// TIA Portal project "TestEssProtoFreia" (V13) (continued)
REGION Network 9: Reset SND_BUSY flag when completed without errors
   RUNG wire#powerrail
      Contact( "SND_DONE(1)" )
      Contact( "SND_BUSY(1)" )
      R_Coil( "SND_BUSY(1)" )
   END_RUNG
   // the same network as SCL:
   IF "SND_DONE(1)" AND "SND_BUSY(1)" THEN "SND_BUSY(1)" := FALSE; END_IF;
END_REGION

REGION Network 10 (STL): Reset SND_BUSY flag and save the status when returned error
         AN    "SND_DONE(1)";
         A     "SND_ERR(1)";
         JNB   ex2;
         R     "SND_BUSY(1)";
         L     "SEND_status(1)";
         T     "SND_STAT_SAVE(1)";
   ex2:  NOP   0;
END_REGION
END_FUNCTION

FUNCTION "Recv_from_Epics" : Void   // FC31, STL
{ S7_Optimized_Access := 'FALSE' }
VERSION : 0.1
BEGIN

REGION Network 1: Get data from Epics (channel 1)
         CALL  AG_RECV
         ( ID     := 1,
           LADDR  := w#16#400,
           RECV   := P#DB101.DBX0.0 BYTE 1000,
           NDR    := "RCV_NDR",
           ERROR  := "RCV_ERR",
           STATUS := "RECV_status",
           LEN    := "RECV_len"
         );
         AN    "RCV_NDR";
         O     "RCV_ERR";
         JC    out;
         CALL  "Cmds_from_Epics";
         BE;
   out:  AN    "RCV_ERR";
         JC    _001;
         L     "RECV_status";
         T     "RCV_STAT_SAVE";
   _001: NOP   0;
END_REGION

REGION Network 2: Get data from Epics (channel 2)
         CALL  AG_RECV
         ( ID     := 2,
           LADDR  := w#16#400,
           RECV   := P#DB105.DBX0.0 BYTE 250,
           NDR    := "RCV_NDR(1)",
           ERROR  := "RCV_ERR(1)",
           STATUS := "RECV_status(1)",
           LEN    := "RECV_len(1)"
         );
         AN    "RCV_NDR(1)";
         O     "RCV_ERR(1)";
         JC    out2;
         CALL  "Data_from_IOC";
         BE;
   out2: AN    "RCV_ERR(1)";
         JC    _002;
         L     "RECV_status(1)";
         T     "RCV_STAT_SAVE(1)";
   _002: NOP   0;
END_REGION
END_FUNCTION

FUNCTION "Send_Epics_data" : Void   // FC32, STL
{ S7_Optimized_Access := 'FALSE' }
VERSION : 0.1
BEGIN

REGION Network 2: Update the Local/remote status
         A     "LocalMode";
         =     "PLC_to_Epics".sLocal;
END_REGION

REGION Network 3: CV01
         L     "CV01_HMI_VAL";
         T     "PLC_to_Epics".CV01.sSetV;
         L     "Tag_7";
         T     "PLC_to_Epics".CV01.sRdV;

         AN    "CV01_ManAuto";
         =     "PLC_to_Epics".CV01.sAuto;
END_REGION

REGION Network 4: CV02
         L     "CV02_HMI_VAL";
         T     "PLC_to_Epics".CV02.sSetV;
         L     "Tag_8";
         T     "PLC_to_Epics".CV02.sRdV;

         AN    "CV02_ManAuto";
         =     "PLC_to_Epics".CV02.sAuto;
END_REGION

REGION Network 5: CV03
         L     "CV03_HMI_VAL";
         T     "PLC_to_Epics".CV03.sSetV;
         L     "Tag_9";
         T     "PLC_to_Epics".CV03.sRdV;

         AN    "CV03_ManAuto";
         =     "PLC_to_Epics".CV03.sAuto;
END_REGION

REGION Network 6: CV04
         L     "CV04_HMI_VAL";
         T     "PLC_to_Epics".CV04.sSetV;
         L     "Tag_10";
         T     "PLC_to_Epics".CV04.sRdV;

         AN    "CV04_ManAuto";
         =     "PLC_to_Epics".CV04.sAuto;
END_REGION

REGION Network 7: CV05
         L     "CV05_HMI_VAL";
         T     "PLC_to_Epics".CV05.sSetV;
         L     "Tag_11";
         T     "PLC_to_Epics".CV05.sRdV;

   //      AN    "CV05_ManAuto"
   //      =     "PLC_to_Epics".CV05.sAuto
END_REGION

REGION Network 8: CV07
         L     "CV07_HMI_VAL";
         T     "PLC_to_Epics".CV07.sSetV;
         L     "Tag_12";
         T     "PLC_to_Epics".CV07.sRdV;

         AN    "CV07_ManAuto";
         =     "PLC_to_Epics".CV07.sAuto;
END_REGION

REGION Network 9: CV60
         L     "CV60_HMI_VAL";
         T     "PLC_to_Epics".CV60.sSetV;
         L     "Tag_13";
         T     "PLC_to_Epics".CV60.sRdV;

         AN    "CV60_ManAuto";
         =     "PLC_to_Epics".CV60.sAuto;
END_REGION

REGION Network 10: CV61
         L     "CV61_HMI_VAL";
         T     "PLC_to_Epics".CV61.sSetV;
         L     "Tag_14";
         T     "PLC_to_Epics".CV61.sRdV;

         AN    "CV61_ManAuto";
         =     "PLC_to_Epics".CV61.sAuto;
END_REGION

REGION Network 11: CV62
         L     "CV62_HMI_VAL";
         T     "PLC_to_Epics".CV62.sSetV;
         L     "Tag_15";
         T     "PLC_to_Epics".CV62.sRdV;

   //      AN    "CV62_ManAuto"
   //      =     "PLC_to_Epics".CV62.sAuto
END_REGION

REGION Network 12: CV550
   //      L     "Tag_14"
   //      T     "PLC_to_Epics".CV550.sRdV

         AN    "ASCOenManuel";
         =     "PLC_to_Epics".CV550.sAuto;
         =     "Data_fo_HNOSS".RegOnMKS2;
END_REGION

REGION Network 13: spare - VB chan 7
         A     "voie 7 chaufferette BV";
         =     "PLC_to_Epics"."spare-VB-7".sHtrOn;
END_REGION

REGION Network 14: spare - VB chan 8
         A     "voie 8 chaufferette BV";
         =     "PLC_to_Epics"."spare-VB-8".sHtrOn;
END_REGION

REGION Network 15: spare VB chan 9
         A     "voie 9 chaufferette BV";
         =     "PLC_to_Epics"."spare-VB-9".sHtrOn;
END_REGION

REGION Network 16: spare - VB chan 10
         A     "voie 10  chaufferette BV";
         =     "PLC_to_Epics"."spare-VB-10".sHtrOn;
END_REGION

REGION Network 17: spare - VB chan 11
         A     "voie 11 chaufferette BV";
         =     "PLC_to_Epics"."spare-VB-11".sHtrOn;
END_REGION

REGION Network 18: EH901-902 CM chan 1
         A     "voie 1 chaufferette CM";
         =     "PLC_to_Epics".EH01.sHtrOn;
END_REGION

REGION Network 19: EH913-914 CM channel 4
         A     "voie 4 chaufferette CM";
         =     "PLC_to_Epics".EH20.sHtrOn;
END_REGION

REGION Network 20: EH933-934 - CM chan 5
         A     "voie 5 chaufferette CM";
         =     "PLC_to_Epics"."spare-CM-5".sHtrOn;
END_REGION

REGION Network 21: EH921 - CM chan 6
         A     "voie 6 chaufferette CM";
         =     "PLC_to_Epics"."spare-CM-6".sHtrOn;
END_REGION

REGION Network 22: EH931-932 - CM chan 7
         A     "voie 7 chaufferette CM";
         =     "PLC_to_Epics"."spare-CM-7".sHtrOn;
END_REGION

REGION Network 23: EH915-916 - CM chan 8
         A     "voie 8 chaufferette CM";
         =     "PLC_to_Epics"."spare-CM-8".sHtrOn;
END_REGION

REGION Network 24: EH937-938 - CM chan 10
         A     "voie 10 chaufferette CM";
         =     "PLC_to_Epics"."spare-CM-10".sHtrOn;
END_REGION

REGION Network 25: EH935-936 - CM chan 12
         A     "voie 12 chaufferette CM";
         =     "PLC_to_Epics"."spare-CM-12".sHtrOn;
END_REGION

REGION Network 26: Status bits
         A     "Graph/manuelle";
         =     "PLC_to_Epics".sManual;
         A     "ErreurSupervision";
         =     "PLC_to_Epics".sGrafcetERR;
         A     "Etat initial";
         =     "PLC_to_Epics".sGS1;
         A     "EtatCdtCryo";
         =     "PLC_to_Epics".sGS2;
         A     "EtatAttMef";
         =     "PLC_to_Epics".sGS3;
         A     "EtatMEFazote";
         =     "PLC_to_Epics".sGS4;
         A     "EtatMEFhelium";
         =     "PLC_to_Epics".sGS5;
         A     "EtatMode4k";
         =     "PLC_to_Epics".sGS6;
         A     "EtatModeStandBy";
         =     "PLC_to_Epics".sGS7;
         A     "EtatMode2K";
         =     "PLC_to_Epics".sGS8;
         A     "Etatrechauffage";
         =     "PLC_to_Epics".sGS10;
         A     "conditionTempMEFheliumOK";
         =     "PLC_to_Epics".sTransTempOK;
         A     "TransMode4K";
         =     "PLC_to_Epics".sTransMode4K;
         A     "EPICS_COMM_OK";
         =     "PLC_to_Epics".EpicsCommOK;
         A     "HNOSS_COMM_OK";
         =     "PLC_to_Epics".HNOSSCommOK;
END_REGION

REGION Network 27: Real parameters read-back (LHe level PID settings)
         L     "TriggerPIDcv01";
         T     "PLC_to_Epics".TrigPID_CV01.sSetV;
         L     "TriggerPIDcv02";
         T     "PLC_to_Epics".TrigPID_CV02.sSetV;
         L     "TriggerPIDcv03";
         T     "PLC_to_Epics".TrigPID_CV03.sSetV;
         L     "LT01LevelSP2k";
         T     "PLC_to_Epics".PID_LT01_CV01_SP.sSetV;
         L     "LT01LevelSP";
         T     "PLC_to_Epics".PID_LT01_CV02_SP.sSetV;
         L     "LT03LevelSP";
         T     "PLC_to_Epics".PID_LT03_CV03_SP.sSetV;
END_REGION

REGION Network 28: Real parameters read-back (CV550l PID settings)
         L     "RéguleASCO02_SP";
         T     "PLC_to_Epics".PID_PT01_CV550_SP.sSetV;
END_REGION

REGION Network 29: Sequence steps
         L     "Data_fo_HNOSS".S4step;
         T     "PLC_to_Epics".S4step;
         L     "Data_fo_HNOSS".S5step;
         T     "PLC_to_Epics".S5step;
         L     "Data_fo_HNOSS".S6step;
         T     "PLC_to_Epics".S6step;
         L     "Data_fo_HNOSS".S7step;
         T     "PLC_to_Epics".S7step;
         L     "Data_fo_HNOSS".S8step;
         T     "PLC_to_Epics".S8step;
         L     "Data_fo_HNOSS".S9step;
         T     "PLC_to_Epics".S9step;
         L     "Data_fo_HNOSS".S10step;
         T     "PLC_to_Epics".S10step;
         L     "Data_fo_HNOSS".SXstep;
         T     "PLC_to_Epics".SXstep;
END_REGION
END_FUNCTION

FUNCTION "Cmds_from_Epics" : Void   // FC33, LAD
TITLE = Process data from Epics
{ S7_Optimized_Access := 'FALSE' }
VERSION : 0.1
   VAR_TEMP   // added for the SCL form of the ladder/FBD networks
      _w1 : Bool;
   END_VAR
BEGIN

REGION Network 1: Switch to remote mode (control from Epics)
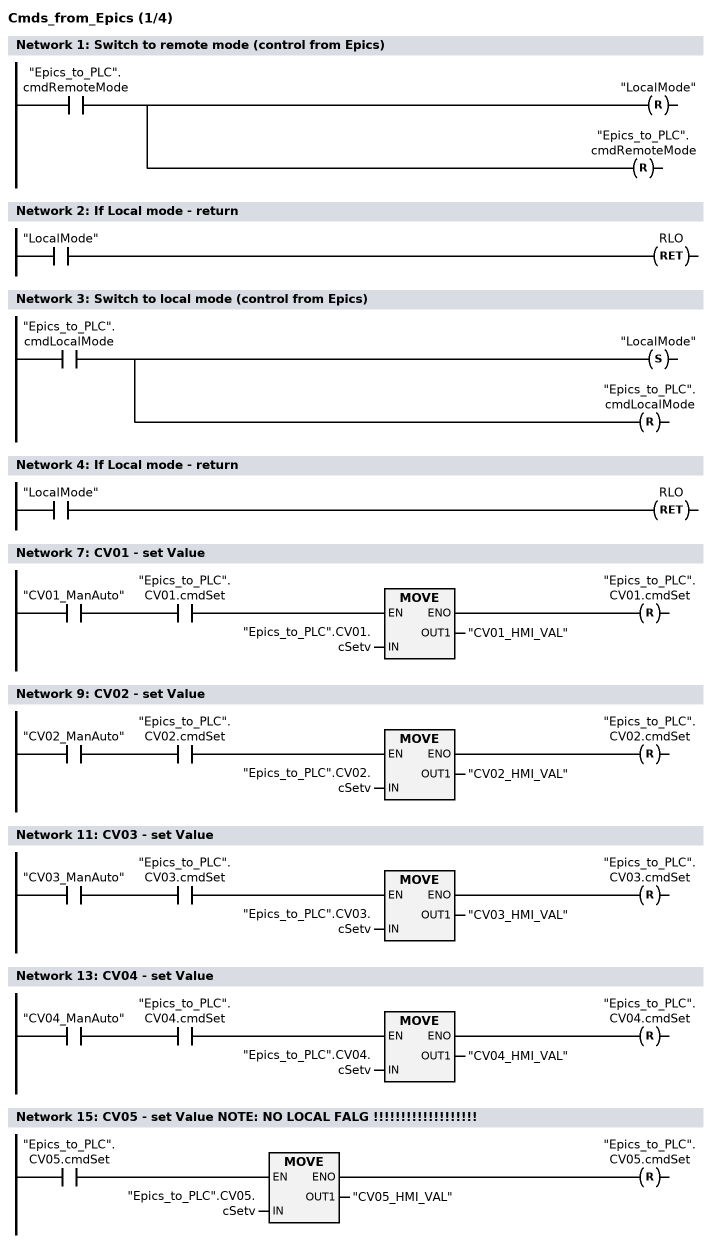
   RUNG wire#powerrail
      Contact( "Epics_to_PLC".cmdRemoteMode )
      wire#w1
      R_Coil( "LocalMode" )
   END_RUNG
   RUNG wire#w1
      R_Coil( "Epics_to_PLC".cmdRemoteMode )
   END_RUNG
   // the same network as SCL:
   IF "Epics_to_PLC".cmdRemoteMode THEN
       "LocalMode" := FALSE;
       "Epics_to_PLC".cmdRemoteMode := FALSE;
   END_IF;
END_REGION

REGION Network 2: If Local mode - return
   IF "LocalMode" THEN
       ENO := TRUE;
       RETURN;
   END_IF;
END_REGION

REGION Network 3: Switch to local mode (control from Epics)
   RUNG wire#powerrail
      Contact( "Epics_to_PLC".cmdLocalMode )
      wire#w1
      S_Coil( "LocalMode" )
   END_RUNG
   RUNG wire#w1
      R_Coil( "Epics_to_PLC".cmdLocalMode )
   END_RUNG
   // the same network as SCL:
   IF "Epics_to_PLC".cmdLocalMode THEN
       "LocalMode" := TRUE;
       "Epics_to_PLC".cmdLocalMode := FALSE;
   END_IF;
END_REGION

REGION Network 4: If Local mode - return
   IF "LocalMode" THEN
       ENO := TRUE;
       RETURN;
   END_IF;
END_REGION

REGION Network 5: Test data (copy block of data)
END_REGION

REGION Network 6 (STL): CV01 Man/Auto
         A     "Epics_to_PLC".CV01.cmdAuto;
         R     "CV01_ManAuto";
         A     "Epics_to_PLC".CV01.cmdMan;
         S     "CV01_ManAuto";
END_REGION

REGION Network 7: CV01 - set Value
   RUNG wire#powerrail
      Contact( "CV01_ManAuto" )
      Contact( "Epics_to_PLC".CV01.cmdSet )
      { S7_GenerateENO := "TRUE" } Move(in := "Epics_to_PLC".CV01.cSetv, out1 => "CV01_HMI_VAL")
      R_Coil( "Epics_to_PLC".CV01.cmdSet )
   END_RUNG
   // the same network as SCL:
   // ENO of a box is taken as its EN; it also drops when the box reports an error
   IF "CV01_ManAuto" AND "Epics_to_PLC".CV01.cmdSet THEN
       "CV01_HMI_VAL" := "Epics_to_PLC".CV01.cSetv;
       "Epics_to_PLC".CV01.cmdSet := FALSE;
   END_IF;
END_REGION

REGION Network 8 (STL): CV02 Man/Auto
         A     "Epics_to_PLC".CV02.cmdAuto;
         R     "CV02_ManAuto";
         A     "Epics_to_PLC".CV02.cmdMan;
         S     "CV02_ManAuto";
END_REGION

REGION Network 9: CV02 - set Value
   RUNG wire#powerrail
      Contact( "CV02_ManAuto" )
      Contact( "Epics_to_PLC".CV02.cmdSet )
      { S7_GenerateENO := "TRUE" } Move(in := "Epics_to_PLC".CV02.cSetv, out1 => "CV02_HMI_VAL")
      R_Coil( "Epics_to_PLC".CV02.cmdSet )
   END_RUNG
   // the same network as SCL:
   // ENO of a box is taken as its EN; it also drops when the box reports an error
   IF "CV02_ManAuto" AND "Epics_to_PLC".CV02.cmdSet THEN
       "CV02_HMI_VAL" := "Epics_to_PLC".CV02.cSetv;
       "Epics_to_PLC".CV02.cmdSet := FALSE;
   END_IF;
END_REGION

REGION Network 10 (STL): CV03 Man/Auto
         A     "Epics_to_PLC".CV03.cmdAuto;
         R     "CV03_ManAuto";
         A     "Epics_to_PLC".CV03.cmdMan;
         S     "CV03_ManAuto";
END_REGION

REGION Network 11: CV03 - set Value
   RUNG wire#powerrail
      Contact( "CV03_ManAuto" )
      Contact( "Epics_to_PLC".CV03.cmdSet )
      { S7_GenerateENO := "TRUE" } Move(in := "Epics_to_PLC".CV03.cSetv, out1 => "CV03_HMI_VAL")
      R_Coil( "Epics_to_PLC".CV03.cmdSet )
   END_RUNG
   // the same network as SCL:
   // ENO of a box is taken as its EN; it also drops when the box reports an error
   IF "CV03_ManAuto" AND "Epics_to_PLC".CV03.cmdSet THEN
       "CV03_HMI_VAL" := "Epics_to_PLC".CV03.cSetv;
       "Epics_to_PLC".CV03.cmdSet := FALSE;
   END_IF;
END_REGION

REGION Network 12 (STL): CV04 Man/Auto
         A     "Epics_to_PLC".CV04.cmdAuto;
         R     "CV04_ManAuto";
         A     "Epics_to_PLC".CV04.cmdMan;
         S     "CV04_ManAuto";
END_REGION

REGION Network 13: CV04 - set Value
   RUNG wire#powerrail
      Contact( "CV04_ManAuto" )
      Contact( "Epics_to_PLC".CV04.cmdSet )
      { S7_GenerateENO := "TRUE" } Move(in := "Epics_to_PLC".CV04.cSetv, out1 => "CV04_HMI_VAL")
      R_Coil( "Epics_to_PLC".CV04.cmdSet )
   END_RUNG
   // the same network as SCL:
   // ENO of a box is taken as its EN; it also drops when the box reports an error
   IF "CV04_ManAuto" AND "Epics_to_PLC".CV04.cmdSet THEN
       "CV04_HMI_VAL" := "Epics_to_PLC".CV04.cSetv;
       "Epics_to_PLC".CV04.cmdSet := FALSE;
   END_IF;
END_REGION

REGION Network 14: CV05 Man/Auto
END_REGION

REGION Network 15: CV05 - set Value NOTE: NO LOCAL FALG !!!!!!!!!!!!!!!!!!!
   RUNG wire#powerrail
      Contact( "Epics_to_PLC".CV05.cmdSet )
      { S7_GenerateENO := "TRUE" } Move(in := "Epics_to_PLC".CV05.cSetv, out1 => "CV05_HMI_VAL")
      R_Coil( "Epics_to_PLC".CV05.cmdSet )
   END_RUNG
   // the same network as SCL:
   // ENO of a box is taken as its EN; it also drops when the box reports an error
   IF "Epics_to_PLC".CV05.cmdSet THEN
       "CV05_HMI_VAL" := "Epics_to_PLC".CV05.cSetv;
       "Epics_to_PLC".CV05.cmdSet := FALSE;
   END_IF;
END_REGION

REGION Network 16 (STL): CV07 Man/Auto
         A     "Epics_to_PLC".CV07.cmdAuto;
         R     "CV07_ManAuto";
         A     "Epics_to_PLC".CV07.cmdMan;
         S     "CV07_ManAuto";
END_REGION

REGION Network 17: CV07 - set Value
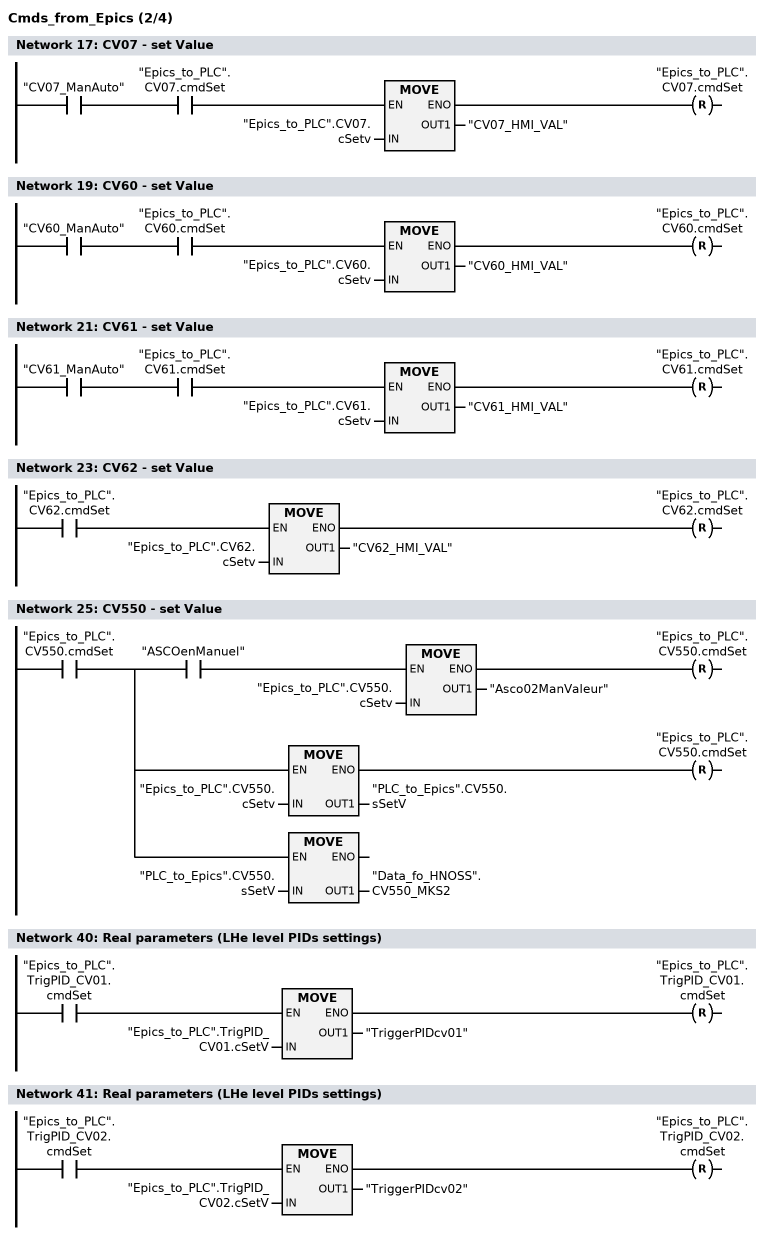
   RUNG wire#powerrail
      Contact( "CV07_ManAuto" )
      Contact( "Epics_to_PLC".CV07.cmdSet )
      { S7_GenerateENO := "TRUE" } Move(in := "Epics_to_PLC".CV07.cSetv, out1 => "CV07_HMI_VAL")
      R_Coil( "Epics_to_PLC".CV07.cmdSet )
   END_RUNG
   // the same network as SCL:
   // ENO of a box is taken as its EN; it also drops when the box reports an error
   IF "CV07_ManAuto" AND "Epics_to_PLC".CV07.cmdSet THEN
       "CV07_HMI_VAL" := "Epics_to_PLC".CV07.cSetv;
       "Epics_to_PLC".CV07.cmdSet := FALSE;
   END_IF;
END_REGION

REGION Network 18 (STL): CV60 Man/Auto
         A     "Epics_to_PLC".CV60.cmdAuto;
         R     "CV60_ManAuto";
         A     "Epics_to_PLC".CV60.cmdMan;
         S     "CV60_ManAuto";
END_REGION

REGION Network 19: CV60 - set Value
   RUNG wire#powerrail
      Contact( "CV60_ManAuto" )
      Contact( "Epics_to_PLC".CV60.cmdSet )
      { S7_GenerateENO := "TRUE" } Move(in := "Epics_to_PLC".CV60.cSetv, out1 => "CV60_HMI_VAL")
      R_Coil( "Epics_to_PLC".CV60.cmdSet )
   END_RUNG
   // the same network as SCL:
   // ENO of a box is taken as its EN; it also drops when the box reports an error
   IF "CV60_ManAuto" AND "Epics_to_PLC".CV60.cmdSet THEN
       "CV60_HMI_VAL" := "Epics_to_PLC".CV60.cSetv;
       "Epics_to_PLC".CV60.cmdSet := FALSE;
   END_IF;
END_REGION

REGION Network 20 (STL): CV61 Man/Auto
         A     "Epics_to_PLC".CV61.cmdAuto;
         R     "CV61_ManAuto";
         A     "Epics_to_PLC".CV61.cmdMan;
         S     "CV61_ManAuto";
END_REGION

REGION Network 21: CV61 - set Value
   RUNG wire#powerrail
      Contact( "CV61_ManAuto" )
      Contact( "Epics_to_PLC".CV61.cmdSet )
      { S7_GenerateENO := "TRUE" } Move(in := "Epics_to_PLC".CV61.cSetv, out1 => "CV61_HMI_VAL")
      R_Coil( "Epics_to_PLC".CV61.cmdSet )
   END_RUNG
   // the same network as SCL:
   // ENO of a box is taken as its EN; it also drops when the box reports an error
   IF "CV61_ManAuto" AND "Epics_to_PLC".CV61.cmdSet THEN
       "CV61_HMI_VAL" := "Epics_to_PLC".CV61.cSetv;
       "Epics_to_PLC".CV61.cmdSet := FALSE;
   END_IF;
END_REGION

REGION Network 22: CV62 Man/Auto
END_REGION

REGION Network 23: CV62 - set Value
   RUNG wire#powerrail
      Contact( "Epics_to_PLC".CV62.cmdSet )
      { S7_GenerateENO := "TRUE" } Move(in := "Epics_to_PLC".CV62.cSetv, out1 => "CV62_HMI_VAL")
      R_Coil( "Epics_to_PLC".CV62.cmdSet )
   END_RUNG
   // the same network as SCL:
   // ENO of a box is taken as its EN; it also drops when the box reports an error
   IF "Epics_to_PLC".CV62.cmdSet THEN
       "CV62_HMI_VAL" := "Epics_to_PLC".CV62.cSetv;
       "Epics_to_PLC".CV62.cmdSet := FALSE;
   END_IF;
END_REGION

REGION Network 24 (STL): CV550 Man/Auto
         A     "Epics_to_PLC".CV550.cmdAuto;
         R     "ASCOenManuel";
         A     "Epics_to_PLC".CV550.cmdMan;
         S     "ASCOenManuel";
END_REGION

REGION Network 25: CV550 - set Value
   RUNG wire#powerrail
      Contact( "Epics_to_PLC".CV550.cmdSet )
      wire#w1
      Contact( "ASCOenManuel" )
      { S7_GenerateENO := "TRUE" } Move(in := "Epics_to_PLC".CV550.cSetv, out1 => "Asco02ManValeur")
      R_Coil( "Epics_to_PLC".CV550.cmdSet )
   END_RUNG
   RUNG wire#w1
      { S7_GenerateENO := "TRUE" } Move(in := "Epics_to_PLC".CV550.cSetv, out1 => "PLC_to_Epics".CV550.sSetV)
      R_Coil( "Epics_to_PLC".CV550.cmdSet )
   END_RUNG
   RUNG wire#w1
      { S7_GenerateENO := "TRUE" } Move(in := "PLC_to_Epics".CV550.sSetV, out1 => "Data_fo_HNOSS".CV550_MKS2)
   END_RUNG
   // the same network as SCL:
   // ENO of a box is taken as its EN; it also drops when the box reports an error
   IF "Epics_to_PLC".CV550.cmdSet AND "ASCOenManuel" THEN
       "Asco02ManValeur" := "Epics_to_PLC".CV550.cSetv;
   END_IF;
   #_w1 := "Epics_to_PLC".CV550.cmdSet;
   IF "Epics_to_PLC".CV550.cmdSet AND "ASCOenManuel" THEN "Epics_to_PLC".CV550.cmdSet := FALSE; END_IF;
   IF #_w1 THEN
       "PLC_to_Epics".CV550.sSetV := "Epics_to_PLC".CV550.cSetv;
       "Epics_to_PLC".CV550.cmdSet := FALSE;
       "Data_fo_HNOSS".CV550_MKS2 := "PLC_to_Epics".CV550.sSetV;
   END_IF;
END_REGION

REGION Network 26 (STL): spare- VB chan 7
         A     "Epics_to_PLC"."spare-VB-7".cmdSet;
         S     "voie 7 chaufferette BV";
         A     "Epics_to_PLC"."spare-VB-7".cmdRst;
         R     "voie 7 chaufferette BV";
END_REGION

REGION Network 27 (STL): spare- VB chan 8
         A     "Epics_to_PLC"."spare-VB-8".cmdSet;
         S     "voie 8 chaufferette BV";
         A     "Epics_to_PLC"."spare-VB-8".cmdRst;
         R     "voie 8 chaufferette BV";
END_REGION

REGION Network 28 (STL): spare- VB chan 9
         A     "Epics_to_PLC"."spare-VB-9".cmdSet;
         S     "voie 9 chaufferette BV";
         A     "Epics_to_PLC"."spare-VB-9".cmdRst;
         R     "voie 9 chaufferette BV";
END_REGION

REGION Network 29 (STL): spare- VB chan 10
         A     "Epics_to_PLC"."spare-VB-10".cmdSet;
         S     "voie 10  chaufferette BV";
         A     "Epics_to_PLC"."spare-VB-10".cmdRst;
         R     "voie 10  chaufferette BV";
END_REGION

REGION Network 30 (STL): spare - VB chan 11
         A     "Epics_to_PLC"."spare-VB-11".cmdSet;
         S     "voie 11 chaufferette BV";
         A     "Epics_to_PLC"."spare-VB-11".cmdRst;
         R     "voie 11 chaufferette BV";
END_REGION

REGION Network 31 (STL): EH901-902 CM chan 1
         A     "Epics_to_PLC".EH01.cmdSet;
         S     "voie 1 chaufferette CM";
         A     "Epics_to_PLC".EH01.cmdRst;
         R     "voie 1 chaufferette CM";
END_REGION

REGION Network 32 (STL): EH913-914 CM chan 4
         A     "Epics_to_PLC".EH20.cmdSet;
         S     "voie 4 chaufferette CM";
         A     "Epics_to_PLC".EH20.cmdRst;
         R     "voie 4 chaufferette CM";
END_REGION

REGION Network 33 (STL): EH933-934 - CM chan 5
         A     "Epics_to_PLC"."spare-CM-5".cmdSet;
         S     "voie 5 chaufferette CM";
         A     "Epics_to_PLC"."spare-CM-5".cmdRst;
         R     "voie 5 chaufferette CM";
END_REGION

REGION Network 34 (STL): EH921 - CM chan 6
         A     "Epics_to_PLC"."spare-CM-6".cmdSet;
         S     "voie 6 chaufferette CM";
         A     "Epics_to_PLC"."spare-CM-6".cmdRst;
         R     "voie 6 chaufferette CM";
END_REGION

REGION Network 35 (STL): EH931-932 - CM chan 7
         A     "Epics_to_PLC"."spare-CM-7".cmdSet;
         S     "voie 7 chaufferette CM";
         A     "Epics_to_PLC"."spare-CM-7".cmdRst;
         R     "voie 7 chaufferette CM";
END_REGION

REGION Network 36 (STL): EH915-916 - CM chan 8
         A     "Epics_to_PLC"."spare-CM-8".cmdSet;
         S     "voie 8 chaufferette CM";
         A     "Epics_to_PLC"."spare-CM-8".cmdRst;
         R     "voie 8 chaufferette CM";
END_REGION

REGION Network 37 (STL): EH937-938 - CM chan 10
         A     "Epics_to_PLC"."spare-CM-10".cmdSet;
         S     "voie 10 chaufferette CM";
         A     "Epics_to_PLC"."spare-CM-10".cmdRst;
         R     "voie 10 chaufferette CM";
END_REGION

REGION Network 38 (STL): EH935-936 - CM chan 12
         A     "Epics_to_PLC"."spare-CM-12".cmdSet;
         S     "voie 12 chaufferette CM";
         A     "Epics_to_PLC"."spare-CM-12".cmdRst;
         R     "voie 12 chaufferette CM";
END_REGION

REGION Network 39 (STL): Bit commands
         A     "Epics_to_PLC".cmdAutoMode;
         R     "Graph/manuelle";
         A     "Epics_to_PLC".cmdManMode;
         S     "Graph/manuelle";
         A     "Epics_to_PLC".cmdGrafcetInit;
         =     "MettreEtatInitial";
         A     "Epics_to_PLC".cmdGrafcetErrRst;
         =     "AcquitterErreurGraph";
         A     "Epics_to_PLC".cmdStartConditioning;
         =     "CmdVanneEtatCdt";
         A     "Epics_to_PLC".cmdCondOK;
         =     "CdtInfraOk";
         A     "Epics_to_PLC".cmdCondERR;
         =     "CdtInfraErreur";
         A     "Epics_to_PLC".cmdStartLN2cooling;
         =     "DmdMefAzote";
         A     "Epics_to_PLC".cmdStartLHecooling;
         =     "DmdMefHelium";
         A     "Epics_to_PLC".cmdStart2Kmode;
         =     "DmdMode2K";
         A     "Epics_to_PLC".cmdStop2Kmode;
         =     "DmdArretMode2k";
         A     "Epics_to_PLC".cmdStartSTBYmode;
         =     "DmdModeStandby";
         A     "Epics_to_PLC".cmdStopSTBYmode;
         =     "DmdArretModeStandby";
         A     "Epics_to_PLC".cmdStartHeating;
         =     "StartHeating";
         A     "Epics_to_PLC".cmdStopHeating;
         =     "StopHeating";
END_REGION

REGION Network 40: Real parameters (LHe level PIDs settings)
   RUNG wire#powerrail
      Contact( "Epics_to_PLC".TrigPID_CV01.cmdSet )
      { S7_GenerateENO := "TRUE" } Move(in := "Epics_to_PLC".TrigPID_CV01.cSetV, out1 => "TriggerPIDcv01")
      R_Coil( "Epics_to_PLC".TrigPID_CV01.cmdSet )
   END_RUNG
   // the same network as SCL:
   // ENO of a box is taken as its EN; it also drops when the box reports an error
   IF "Epics_to_PLC".TrigPID_CV01.cmdSet THEN
       "TriggerPIDcv01" := "Epics_to_PLC".TrigPID_CV01.cSetV;
       "Epics_to_PLC".TrigPID_CV01.cmdSet := FALSE;
   END_IF;
END_REGION

REGION Network 41: Real parameters (LHe level PIDs settings)
   RUNG wire#powerrail
      Contact( "Epics_to_PLC".TrigPID_CV02.cmdSet )
      { S7_GenerateENO := "TRUE" } Move(in := "Epics_to_PLC".TrigPID_CV02.cSetV, out1 => "TriggerPIDcv02")
      R_Coil( "Epics_to_PLC".TrigPID_CV02.cmdSet )
   END_RUNG
   // the same network as SCL:
   // ENO of a box is taken as its EN; it also drops when the box reports an error
   IF "Epics_to_PLC".TrigPID_CV02.cmdSet THEN
       "TriggerPIDcv02" := "Epics_to_PLC".TrigPID_CV02.cSetV;
       "Epics_to_PLC".TrigPID_CV02.cmdSet := FALSE;
   END_IF;
END_REGION

REGION Network 42: Real parameters (LHe level PIDs settings)
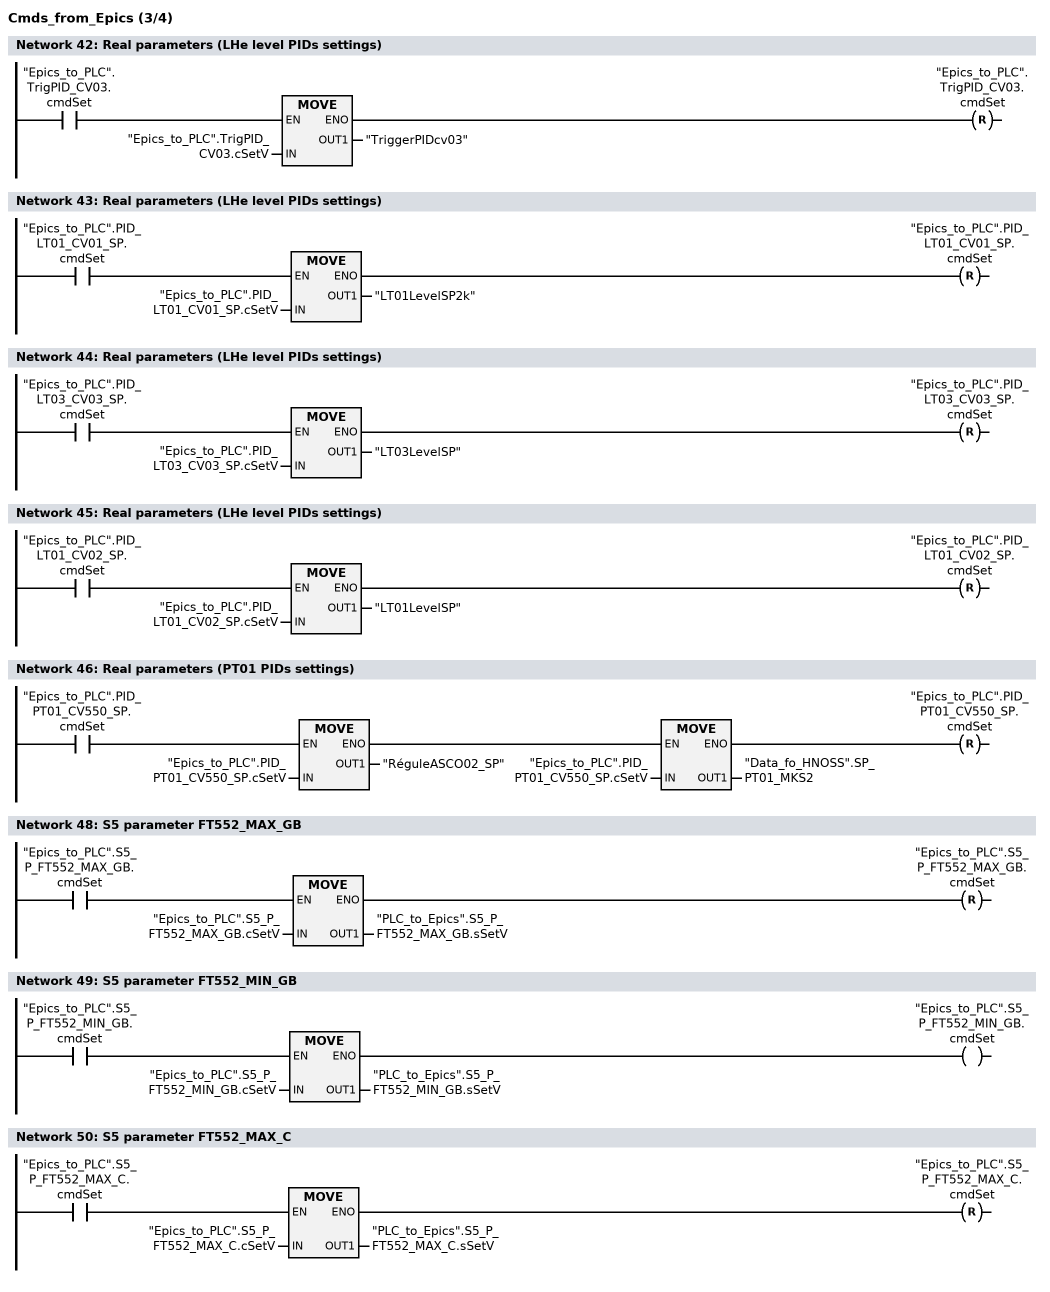
   RUNG wire#powerrail
      Contact( "Epics_to_PLC".TrigPID_CV03.cmdSet )
      { S7_GenerateENO := "TRUE" } Move(in := "Epics_to_PLC".TrigPID_CV03.cSetV, out1 => "TriggerPIDcv03")
      R_Coil( "Epics_to_PLC".TrigPID_CV03.cmdSet )
   END_RUNG
   // the same network as SCL:
   // ENO of a box is taken as its EN; it also drops when the box reports an error
   IF "Epics_to_PLC".TrigPID_CV03.cmdSet THEN
       "TriggerPIDcv03" := "Epics_to_PLC".TrigPID_CV03.cSetV;
       "Epics_to_PLC".TrigPID_CV03.cmdSet := FALSE;
   END_IF;
END_REGION

REGION Network 43: Real parameters (LHe level PIDs settings)
   RUNG wire#powerrail
      Contact( "Epics_to_PLC".PID_LT01_CV01_SP.cmdSet )
      { S7_GenerateENO := "TRUE" } Move(in := "Epics_to_PLC".PID_LT01_CV01_SP.cSetV, out1 => "LT01LevelSP2k")
      R_Coil( "Epics_to_PLC".PID_LT01_CV01_SP.cmdSet )
   END_RUNG
   // the same network as SCL:
   // ENO of a box is taken as its EN; it also drops when the box reports an error
   IF "Epics_to_PLC".PID_LT01_CV01_SP.cmdSet THEN
       "LT01LevelSP2k" := "Epics_to_PLC".PID_LT01_CV01_SP.cSetV;
       "Epics_to_PLC".PID_LT01_CV01_SP.cmdSet := FALSE;
   END_IF;
END_REGION

REGION Network 44: Real parameters (LHe level PIDs settings)
   RUNG wire#powerrail
      Contact( "Epics_to_PLC".PID_LT03_CV03_SP.cmdSet )
      { S7_GenerateENO := "TRUE" } Move(in := "Epics_to_PLC".PID_LT03_CV03_SP.cSetV, out1 => "LT03LevelSP")
      R_Coil( "Epics_to_PLC".PID_LT03_CV03_SP.cmdSet )
   END_RUNG
   // the same network as SCL:
   // ENO of a box is taken as its EN; it also drops when the box reports an error
   IF "Epics_to_PLC".PID_LT03_CV03_SP.cmdSet THEN
       "LT03LevelSP" := "Epics_to_PLC".PID_LT03_CV03_SP.cSetV;
       "Epics_to_PLC".PID_LT03_CV03_SP.cmdSet := FALSE;
   END_IF;
END_REGION

REGION Network 45: Real parameters (LHe level PIDs settings)
   RUNG wire#powerrail
      Contact( "Epics_to_PLC".PID_LT01_CV02_SP.cmdSet )
      { S7_GenerateENO := "TRUE" } Move(in := "Epics_to_PLC".PID_LT01_CV02_SP.cSetV, out1 => "LT01LevelSP")
      R_Coil( "Epics_to_PLC".PID_LT01_CV02_SP.cmdSet )
   END_RUNG
   // the same network as SCL:
   // ENO of a box is taken as its EN; it also drops when the box reports an error
   IF "Epics_to_PLC".PID_LT01_CV02_SP.cmdSet THEN
       "LT01LevelSP" := "Epics_to_PLC".PID_LT01_CV02_SP.cSetV;
       "Epics_to_PLC".PID_LT01_CV02_SP.cmdSet := FALSE;
   END_IF;
END_REGION

REGION Network 46: Real parameters (PT01 PIDs settings)
   RUNG wire#powerrail
      Contact( "Epics_to_PLC".PID_PT01_CV550_SP.cmdSet )
      { S7_GenerateENO := "TRUE" } Move(in := "Epics_to_PLC".PID_PT01_CV550_SP.cSetV, out1 => "RéguleASCO02_SP")
      { S7_GenerateENO := "TRUE" } Move(in := "Epics_to_PLC".PID_PT01_CV550_SP.cSetV, out1 => "Data_fo_HNOSS".SP_PT01_MKS2)
      R_Coil( "Epics_to_PLC".PID_PT01_CV550_SP.cmdSet )
   END_RUNG
   // the same network as SCL:
   // ENO of a box is taken as its EN; it also drops when the box reports an error
   IF "Epics_to_PLC".PID_PT01_CV550_SP.cmdSet THEN
       "RéguleASCO02_SP" := "Epics_to_PLC".PID_PT01_CV550_SP.cSetV;
       "Data_fo_HNOSS".SP_PT01_MKS2 := "Epics_to_PLC".PID_PT01_CV550_SP.cSetV;
       "Epics_to_PLC".PID_PT01_CV550_SP.cmdSet := FALSE;
   END_IF;
END_REGION

REGION Network 47 (STL): Temperatures fromKeithley
         L     "Epics_to_PLC".TTxx;
         T     "ReceivePT100"."TTxx_(K)";
         L     "Epics_to_PLC".TTyy;
         T     "ReceivePT100"."TTyy_(K)";
END_REGION

REGION Network 48: S5 parameter FT552_MAX_GB
   RUNG wire#powerrail
      Contact( "Epics_to_PLC".S5_P_FT552_MAX_GB.cmdSet )
      { S7_GenerateENO := "TRUE" } Move(in := "Epics_to_PLC".S5_P_FT552_MAX_GB.cSetV, out1 => "PLC_to_Epics".S5_P_FT552_MAX_GB.sSetV)
      R_Coil( "Epics_to_PLC".S5_P_FT552_MAX_GB.cmdSet )
   END_RUNG
   // the same network as SCL:
   // ENO of a box is taken as its EN; it also drops when the box reports an error
   IF "Epics_to_PLC".S5_P_FT552_MAX_GB.cmdSet THEN
       "PLC_to_Epics".S5_P_FT552_MAX_GB.sSetV := "Epics_to_PLC".S5_P_FT552_MAX_GB.cSetV;
       "Epics_to_PLC".S5_P_FT552_MAX_GB.cmdSet := FALSE;
   END_IF;
END_REGION

REGION Network 49: S5 parameter FT552_MIN_GB
   RUNG wire#powerrail
      Contact( "Epics_to_PLC".S5_P_FT552_MIN_GB.cmdSet )
      { S7_GenerateENO := "TRUE" } Move(in := "Epics_to_PLC".S5_P_FT552_MIN_GB.cSetV, out1 => "PLC_to_Epics".S5_P_FT552_MIN_GB.sSetV)
      Coil( "Epics_to_PLC".S5_P_FT552_MIN_GB.cmdSet )
   END_RUNG
   // the same network as SCL:
   // ENO of a box is taken as its EN; it also drops when the box reports an error
   IF "Epics_to_PLC".S5_P_FT552_MIN_GB.cmdSet THEN
       "PLC_to_Epics".S5_P_FT552_MIN_GB.sSetV := "Epics_to_PLC".S5_P_FT552_MIN_GB.cSetV;
   END_IF;
   "Epics_to_PLC".S5_P_FT552_MIN_GB.cmdSet := "Epics_to_PLC".S5_P_FT552_MIN_GB.cmdSet;
END_REGION

REGION Network 50: S5 parameter FT552_MAX_C
   RUNG wire#powerrail
      Contact( "Epics_to_PLC".S5_P_FT552_MAX_C.cmdSet )
      { S7_GenerateENO := "TRUE" } Move(in := "Epics_to_PLC".S5_P_FT552_MAX_C.cSetV, out1 => "PLC_to_Epics".S5_P_FT552_MAX_C.sSetV)
      R_Coil( "Epics_to_PLC".S5_P_FT552_MAX_C.cmdSet )
   END_RUNG
   // the same network as SCL:
   // ENO of a box is taken as its EN; it also drops when the box reports an error
   IF "Epics_to_PLC".S5_P_FT552_MAX_C.cmdSet THEN
       "PLC_to_Epics".S5_P_FT552_MAX_C.sSetV := "Epics_to_PLC".S5_P_FT552_MAX_C.cSetV;
       "Epics_to_PLC".S5_P_FT552_MAX_C.cmdSet := FALSE;
   END_IF;
END_REGION

REGION Network 51: S5 parameter FT552_MIN_C
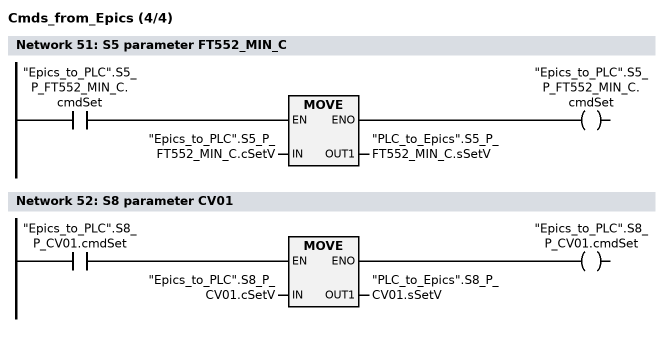
   RUNG wire#powerrail
      Contact( "Epics_to_PLC".S5_P_FT552_MIN_C.cmdSet )
      { S7_GenerateENO := "TRUE" } Move(in := "Epics_to_PLC".S5_P_FT552_MIN_C.cSetV, out1 => "PLC_to_Epics".S5_P_FT552_MIN_C.sSetV)
      Coil( "Epics_to_PLC".S5_P_FT552_MIN_C.cmdSet )
   END_RUNG
   // the same network as SCL:
   // ENO of a box is taken as its EN; it also drops when the box reports an error
   IF "Epics_to_PLC".S5_P_FT552_MIN_C.cmdSet THEN
       "PLC_to_Epics".S5_P_FT552_MIN_C.sSetV := "Epics_to_PLC".S5_P_FT552_MIN_C.cSetV;
   END_IF;
   "Epics_to_PLC".S5_P_FT552_MIN_C.cmdSet := "Epics_to_PLC".S5_P_FT552_MIN_C.cmdSet;
END_REGION

REGION Network 52: S8 parameter CV01
   RUNG wire#powerrail
      Contact( "Epics_to_PLC".S8_P_CV01.cmdSet )
      { S7_GenerateENO := "TRUE" } Move(in := "Epics_to_PLC".S8_P_CV01.cSetV, out1 => "PLC_to_Epics".S8_P_CV01.sSetV)
      Coil( "Epics_to_PLC".S8_P_CV01.cmdSet )
   END_RUNG
   // the same network as SCL:
   // ENO of a box is taken as its EN; it also drops when the box reports an error
   IF "Epics_to_PLC".S8_P_CV01.cmdSet THEN
       "PLC_to_Epics".S8_P_CV01.sSetV := "Epics_to_PLC".S8_P_CV01.cSetV;
   END_IF;
   "Epics_to_PLC".S8_P_CV01.cmdSet := "Epics_to_PLC".S8_P_CV01.cmdSet;
END_REGION
END_FUNCTION

FUNCTION "Data_from_IOC" : Void   // FC34, LAD
TITLE = Get data from the IOC andcheck if the connection is alive
{ S7_Optimized_Access := 'FALSE' }
VERSION : 0.1
BEGIN

REGION Network 1: Check the Data from the IOC
END_REGION
END_FUNCTION

FUNCTION "grafcet" : Void   // FC99, LAD
{ S7_Optimized_Access := 'FALSE' }
VERSION : 0.1
   VAR_TEMP   // added for the SCL form of the ladder/FBD networks
      _w1 : Bool;
      _w2 : Bool;
      _w3 : Bool;
      _w4 : Bool;
      _w5 : Bool;
      _w6 : Bool;
      _w7 : Bool;
      _w8 : Bool;
   END_VAR
BEGIN

REGION Network 1: Set initial step number for the state S4
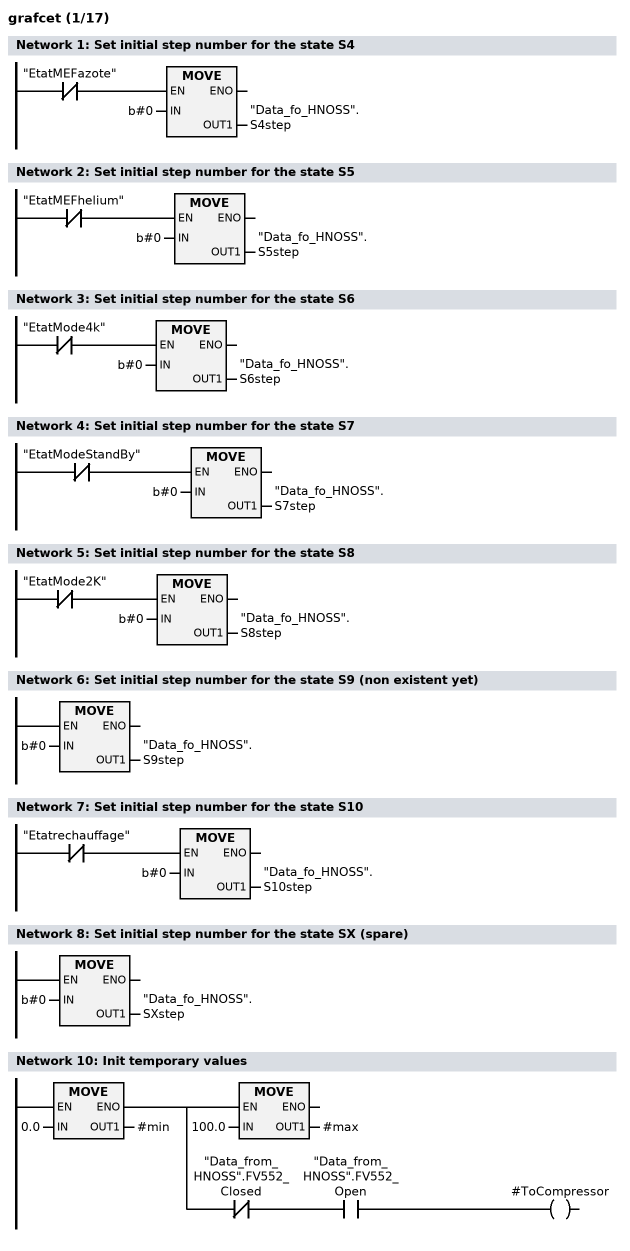
   RUNG wire#powerrail
      I_Contact( "EtatMEFazote" )
      { S7_GenerateENO := "TRUE" } Move(in := b#0, out1 => "Data_fo_HNOSS".S4step)
   END_RUNG
   // the same network as SCL:
   IF NOT "EtatMEFazote" THEN "Data_fo_HNOSS".S4step := b#0; END_IF;
END_REGION

